// TIA Portal project "Catalyst_syzygy_v2.1" (V17) (continued)
VERSION : 1.0
// stored: InstanceOfName TX-AI
"TX-AI"
BEGIN
   Retain.HMI.Config.ESMXV := 50.0;
   Retain.HMI.Config.SP.Limits.H := 10.0;
   Retain.HMI.Config.SP.Limits.HH := 50.0;
END_DATA_BLOCK

// folder: Analogs inputs/Trasmitters/Level Trasmitters/Datablocks

DATA_BLOCK "LT-1011_DB"   // DB8
{ S7_Optimized_Access := 'TRUE' }
VERSION : 1.0
// stored: InstanceOfName TX-AI
"TX-AI"
BEGIN
   Retain.HMI.Config.SP.Limits.H := 85.0;
   Retain.HMI.Config.SP.Limits.HH := 95.0;
END_DATA_BLOCK

DATA_BLOCK "LT-1061_DB"   // DB9
{ S7_Optimized_Access := 'TRUE' }
VERSION : 1.0
// stored: InstanceOfName TX-AI
"TX-AI"
BEGIN
END_DATA_BLOCK

DATA_BLOCK "LT-1021_DB"   // DB35
{ S7_Optimized_Access := 'TRUE' }
VERSION : 1.0
// stored: InstanceOfName TX-AI
"TX-AI"
BEGIN
END_DATA_BLOCK

DATA_BLOCK "LT-2011_DB"   // DB49
{ S7_Optimized_Access := 'TRUE' }
VERSION : 1.0
// stored: InstanceOfName TX-AI
"TX-AI"
BEGIN
   Retain.HMI.Config.SP.Limits.L := 18.0;
END_DATA_BLOCK

DATA_BLOCK "LT-2021_DB"   // DB56
{ S7_Optimized_Access := 'TRUE' }
VERSION : 1.0
// stored: InstanceOfName TX-AI
"TX-AI"
BEGIN
   Retain.HMI.Config.SP.Limits.L := 18.0;
END_DATA_BLOCK

DATA_BLOCK "LT-1031_DB"   // DB60
{ S7_Optimized_Access := 'TRUE' }
VERSION : 1.0
// stored: InstanceOfName TX-AI
"TX-AI"
BEGIN
END_DATA_BLOCK

DATA_BLOCK "LT-1051_DB"   // DB120
{ S7_Optimized_Access := 'TRUE' }
VERSION : 1.0
// stored: InstanceOfName TX-AI
"TX-AI"
BEGIN
END_DATA_BLOCK

DATA_BLOCK "LT-1011_VOL_DB"   // DB152
{ S7_Optimized_Access := 'TRUE' }
VERSION : 1.0
// stored: InstanceOfName TX-AI
"TX-AI"
BEGIN
   Retain.HMI.Config.ESMXV := 1133.72;
   Retain.HMI.Config.SP.Limits.H := 1000.0;
   Retain.HMI.Config.SP.Limits.HH := 1100.0;
END_DATA_BLOCK

DATA_BLOCK "LT-1061_VOL_DB"   // DB232
{ S7_Optimized_Access := 'TRUE' }
VERSION : 1.0
// stored: InstanceOfName TX-AI
"TX-AI"
BEGIN
END_DATA_BLOCK

DATA_BLOCK "LT-1021_VOL_DB"   // DB243
{ S7_Optimized_Access := 'TRUE' }
VERSION : 1.0
// stored: InstanceOfName TX-AI
"TX-AI"
BEGIN
   Retain.HMI.Config.ESMXV := 2300.0;
   Retain.HMI.Config.SP.Limits.H := 2000.0;
   Retain.HMI.Config.SP.Limits.HH := 2100.0;
END_DATA_BLOCK

DATA_BLOCK "LT-1031_VOL_DB"   // DB245
{ S7_Optimized_Access := 'TRUE' }
VERSION : 1.0
// stored: InstanceOfName TX-AI
"TX-AI"
BEGIN
   Retain.HMI.Config.ESMXV := 500.0;
   Retain.HMI.Config.SP.Limits.H := 450.0;
   Retain.HMI.Config.SP.Limits.HH := 480.0;
END_DATA_BLOCK

DATA_BLOCK "LT-1051_VOL_DB"   // DB246
{ S7_Optimized_Access := 'TRUE' }
VERSION : 1.0
// stored: InstanceOfName TX-AI
"TX-AI"
BEGIN
END_DATA_BLOCK

DATA_BLOCK "LT-2011_VOL_DB"   // DB247
{ S7_Optimized_Access := 'TRUE' }
VERSION : 1.0
// stored: InstanceOfName TX-AI
"TX-AI"
BEGIN
   Retain.HMI.Config.ESMXV := 200.0;
   Retain.HMI.Config.SP.Limits.H := 180.0;
   Retain.HMI.Config.SP.Limits.HH := 190.0;
END_DATA_BLOCK

DATA_BLOCK "LT-2021_VOL_DB"   // DB248
{ S7_Optimized_Access := 'TRUE' }
VERSION : 1.0
// stored: InstanceOfName TX-AI
"TX-AI"
BEGIN
   Retain.HMI.Config.ESMXV := 200.0;
   Retain.HMI.Config.SP.Limits.H := 180.0;
   Retain.HMI.Config.SP.Limits.HH := 190.0;
END_DATA_BLOCK

// folder: Analogs inputs/Trasmitters/Ph Trasmitters/Datablocks

DATA_BLOCK "pH-2011_DB"   // DB46
{ S7_Optimized_Access := 'TRUE' }
VERSION : 1.0
// stored: InstanceOfName TX-AI
"TX-AI"
BEGIN
   Retain.HMI.Config.ESMXV := 14.0;
   Retain.HMI.Config.SP.Limits.HH := 12.0;
   Retain.HMI.Config.SP.Limits.H := 10.0;
END_DATA_BLOCK

DATA_BLOCK "pH-2012_DB"   // DB47
{ S7_Optimized_Access := 'TRUE' }
VERSION : 1.0
// stored: InstanceOfName TX-AI
"TX-AI"
BEGIN
   Retain.HMI.Config.ESMXV := 14.0;
   Retain.HMI.Config.SP.Limits.HH := 12.0;
   Retain.HMI.Config.SP.Limits.H := 10.0;
END_DATA_BLOCK

DATA_BLOCK "pH-2021_DB"   // DB54
{ S7_Optimized_Access := 'TRUE' }
VERSION : 1.0
// stored: InstanceOfName TX-AI
"TX-AI"
BEGIN
   Retain.HMI.Config.ESMXV := 14.0;
   Retain.HMI.Config.SP.Limits.HH := 12.0;
   Retain.HMI.Config.SP.Limits.H := 10.0;
END_DATA_BLOCK

DATA_BLOCK "pH-2022_DB"   // DB55
{ S7_Optimized_Access := 'TRUE' }
VERSION : 1.0
// stored: InstanceOfName TX-AI
"TX-AI"
BEGIN
   Retain.HMI.Config.ESMXV := 14.0;
   Retain.HMI.Config.SP.Limits.HH := 12.0;
   Retain.HMI.Config.SP.Limits.H := 10.0;
END_DATA_BLOCK

// folder: Analogs inputs/Trasmitters/Pressure Trasmitters/Datablocks

DATA_BLOCK "PT-101A_DB"   // DB31
{ S7_Optimized_Access := 'TRUE' }
VERSION : 1.0
// stored: InstanceOfName TX-AI
"TX-AI"
BEGIN
   Retain.HMI.Config.SP.Limits.HH := 124.0;
   Retain.HMI.Config.SP.Limits.H := 120.0;
   Retain.HMI.Config.ESMXV := 125.0;
END_DATA_BLOCK

DATA_BLOCK "PT-101B_DB"   // DB32
{ S7_Optimized_Access := 'TRUE' }
VERSION : 1.0
// stored: InstanceOfName TX-AI
"TX-AI"
BEGIN
   Retain.HMI.Config.SP.Limits.HH := 124.0;
   Retain.HMI.Config.SP.Limits.H := 120.0;
   Retain.HMI.Config.ESMXV := 125.0;
END_DATA_BLOCK

DATA_BLOCK "PT-102A_DB"   // DB36
{ S7_Optimized_Access := 'TRUE' }
VERSION : 1.0
// stored: InstanceOfName TX-AI
"TX-AI"
BEGIN
   Retain.HMI.Config.ESMXV := 125.0;
   Retain.HMI.Config.SP.Limits.HH := 124.0;
   Retain.HMI.Config.SP.Limits.H := 120.0;
END_DATA_BLOCK

DATA_BLOCK "PT-102B_DB"   // DB37
{ S7_Optimized_Access := 'TRUE' }
VERSION : 1.0
// stored: InstanceOfName TX-AI
"TX-AI"
BEGIN
   Retain.HMI.Config.ESMXV := 125.0;
   Retain.HMI.Config.SP.Limits.HH := 124.0;
   Retain.HMI.Config.SP.Limits.H := 120.0;
END_DATA_BLOCK

DATA_BLOCK "PT-201A_DB"   // DB50
{ S7_Optimized_Access := 'TRUE' }
VERSION : 1.0
// stored: InstanceOfName TX-AI
"TX-AI"
BEGIN
   Retain.HMI.Config.ESMXV := 125.0;
   Retain.HMI.Config.SP.Limits.HH := 110.0;
   Retain.HMI.Config.SP.Limits.H := 100.0;
END_DATA_BLOCK

DATA_BLOCK "PT-201B_DB"   // DB51
{ S7_Optimized_Access := 'TRUE' }
VERSION : 1.0
// stored: InstanceOfName TX-AI
"TX-AI"
BEGIN
   Retain.HMI.Config.ESMXV := 125.0;
   Retain.HMI.Config.SP.Limits.HH := 110.0;
   Retain.HMI.Config.SP.Limits.H := 100.0;
END_DATA_BLOCK

DATA_BLOCK "PT-202A_DB"   // DB57
{ S7_Optimized_Access := 'TRUE' }
VERSION : 1.0
// stored: InstanceOfName TX-AI
"TX-AI"
BEGIN
   Retain.HMI.Config.ESMXV := 125.0;
   Retain.HMI.Config.SP.Limits.HH := 110.0;
   Retain.HMI.Config.SP.Limits.H := 100.0;
END_DATA_BLOCK

DATA_BLOCK "PT-202B_DB"   // DB58
{ S7_Optimized_Access := 'TRUE' }
VERSION : 1.0
// stored: InstanceOfName TX-AI
"TX-AI"
BEGIN
   Retain.HMI.Config.ESMXV := 125.0;
   Retain.HMI.Config.SP.Limits.HH := 110.0;
   Retain.HMI.Config.SP.Limits.H := 100.0;
END_DATA_BLOCK

DATA_BLOCK "PT-103A_DB"   // DB61
{ S7_Optimized_Access := 'TRUE' }
VERSION : 1.0
// stored: InstanceOfName TX-AI
"TX-AI"
BEGIN
   Retain.HMI.Config.ESMXV := 125.0;
   Retain.HMI.Config.SP.Limits.H := 124.0;
   Retain.HMI.Config.SP.Limits.L := 120.0;
END_DATA_BLOCK

DATA_BLOCK "PT-103B_DB"   // DB62
{ S7_Optimized_Access := 'TRUE' }
VERSION : 1.0
// stored: InstanceOfName TX-AI
"TX-AI"
BEGIN
   Retain.HMI.Config.ESMXV := 125.0;
   Retain.HMI.Config.SP.Limits.HH := 124.0;
   Retain.HMI.Config.SP.Limits.H := 120.0;
END_DATA_BLOCK

DATA_BLOCK "PT-301A_DB"   // DB64
{ S7_Optimized_Access := 'TRUE' }
VERSION : 1.0
// stored: InstanceOfName TX-AI
"TX-AI"
BEGIN
   Retain.HMI.Config.ESMXV := 125.0;
   Retain.HMI.Config.SP.Limits.HH := 110.0;
   Retain.HMI.Config.SP.Limits.H := 100.0;
END_DATA_BLOCK

DATA_BLOCK "PT-301B_DB"   // DB65
{ S7_Optimized_Access := 'TRUE' }
VERSION : 1.0
// stored: InstanceOfName TX-AI
"TX-AI"
BEGIN
   Retain.HMI.Config.ESMXV := 125.0;
   Retain.HMI.Config.SP.Limits.HH := 110.0;
   Retain.HMI.Config.SP.Limits.H := 100.0;
END_DATA_BLOCK

DATA_BLOCK "PT-104A_DB"   // DB124
{ S7_Optimized_Access := 'TRUE' }
VERSION : 1.0
// stored: InstanceOfName TX-AI
"TX-AI"
BEGIN
   Retain.HMI.Config.ESMXV := 64.0;
END_DATA_BLOCK

DATA_BLOCK "PT-104B_DB"   // DB125
{ S7_Optimized_Access := 'TRUE' }
VERSION : 1.0
// stored: InstanceOfName TX-AI
"TX-AI"
BEGIN
   Retain.HMI.Config.ESMXV := 64.0;
END_DATA_BLOCK

DATA_BLOCK "MFC-4011-P_DB"   // DB162
{ S7_Optimized_Access := 'TRUE' }
VERSION : 1.0
// stored: InstanceOfName TX-AI
"TX-AI"
BEGIN
   Retain.HMI.Config.SP.Limits.HH := 17.3;
   Retain.HMI.Config.SP.Limits.H := 16.3;
   Retain.HMI.Config.SP.Limits.L := 15.0;
   Retain.HMI.Config.SP.Limits.LL := 14.8;
   Retain.HMI.Config.PT.HLD.ALL := t#15s;
   Retain.HMI.Config.PT.HLD.AHH := t#15s;
END_DATA_BLOCK

DATA_BLOCK "PT-M_4024_DB"   // DB165
{ S7_Optimized_Access := 'TRUE' }
VERSION : 1.0
// stored: InstanceOfName TX-AI
"TX-AI"
BEGIN
END_DATA_BLOCK

DATA_BLOCK "PT-M_4025_DB"   // DB166
{ S7_Optimized_Access := 'TRUE' }
VERSION : 1.0
// stored: InstanceOfName TX-AI
"TX-AI"
BEGIN
END_DATA_BLOCK

DATA_BLOCK "MFC-4012-P_DB"   // DB176
{ S7_Optimized_Access := 'TRUE' }
VERSION : 1.0
// stored: InstanceOfName TX-AI
"TX-AI"
BEGIN
END_DATA_BLOCK

DATA_BLOCK "MFC-4024-P_DB"   // DB213
{ S7_Optimized_Access := 'TRUE' }
VERSION : 1.0
// stored: InstanceOfName TX-AI
"TX-AI"
BEGIN
END_DATA_BLOCK

DATA_BLOCK "MFC-4025-P_DB"   // DB216
{ S7_Optimized_Access := 'TRUE' }
VERSION : 1.0
// stored: InstanceOfName TX-AI
"TX-AI"
BEGIN
END_DATA_BLOCK

DATA_BLOCK "MFC-4021-P_DB"   // DB398
{ S7_Optimized_Access := 'TRUE' }
VERSION : 1.0
// stored: InstanceOfName TX-AI
"TX-AI"
BEGIN
END_DATA_BLOCK

// folder: Analogs inputs/Trasmitters/Temperature Trasmitters/DataBlocks

DATA_BLOCK "TT-2011_DB"   // DB44
{ S7_Optimized_Access := 'TRUE' }
VERSION : 1.0
// stored: InstanceOfName TX-AI
"TX-AI"
BEGIN
   Retain.HMI.Config.SP.Limits.L := 75.0;
   Retain.HMI.Config.SP.Limits.LL := 70.0;
   Retain.HMI.Config.ESMXV := 200.0;
END_DATA_BLOCK

DATA_BLOCK "TT-2012_DB"   // DB45
{ S7_Optimized_Access := 'TRUE' }
VERSION : 1.0
// stored: InstanceOfName TX-AI
"TX-AI"
BEGIN
   Retain.HMI.Config.SP.Limits.L := 75.0;
   Retain.HMI.Config.SP.Limits.LL := 70.0;
   Retain.HMI.Config.ESMXV := 200.0;
END_DATA_BLOCK

DATA_BLOCK "TT-2021_DB"   // DB52
{ S7_Optimized_Access := 'TRUE' }
VERSION : 1.0
// stored: InstanceOfName TX-AI
"TX-AI"
BEGIN
   Retain.HMI.Config.ESMXV := 200.0;
   Retain.HMI.Config.SP.Limits.L := 70.0;
   Retain.HMI.Config.SP.Limits.LL := 75.0;
END_DATA_BLOCK

DATA_BLOCK "TT-2022_DB"   // DB53
{ S7_Optimized_Access := 'TRUE' }
VERSION : 1.0
// stored: InstanceOfName TX-AI
"TX-AI"
BEGIN
   Retain.HMI.Config.SP.Limits.L := 75.0;
   Retain.HMI.Config.SP.Limits.LL := 70.0;
   Retain.HMI.Config.ESMXV := 200.0;
END_DATA_BLOCK

DATA_BLOCK "TT-1031_DB"   // DB59
{ S7_Optimized_Access := 'TRUE' }
VERSION : 1.0
// stored: InstanceOfName TX-AI
"TX-AI"
BEGIN
   Retain.HMI.Config.ESMXV := 200.0;
END_DATA_BLOCK

DATA_BLOCK "TT-401A_DB"   // DB69
{ S7_Optimized_Access := 'TRUE' }
VERSION : 1.0
// stored: InstanceOfName TX-AI
"TX-AI"
BEGIN
   Retain.HMI.Config.ESMXV := 1350.0;
   Retain.HMI.Config.RIMXV := 13500.0;
   Retain.HMI.Config.SP.Limits.HH := 800.0;
   Retain.HMI.Config.SP.Limits.H := 750.0;
END_DATA_BLOCK

DATA_BLOCK "TT-401B_DB"   // DB70
{ S7_Optimized_Access := 'TRUE' }
VERSION : 1.0
// stored: InstanceOfName TX-AI
"TX-AI"
BEGIN
   Retain.HMI.Config.ESMXV := 1350.0;
   Retain.HMI.Config.RIMXV := 13500.0;
   Retain.HMI.Config.SP.Limits.HH := 800.0;
   Retain.HMI.Config.SP.Limits.H := 750.0;
END_DATA_BLOCK

DATA_BLOCK "TT-401C_DB"   // DB71
{ S7_Optimized_Access := 'TRUE' }
VERSION : 1.0
// stored: InstanceOfName TX-AI
"TX-AI"
BEGIN
   Retain.HMI.Config.ESMXV := 1350.0;
   Retain.HMI.Config.RIMXV := 13500.0;
   Retain.HMI.Config.SP.Limits.HH := 800.0;
   Retain.HMI.Config.SP.Limits.H := 750.0;
END_DATA_BLOCK

DATA_BLOCK "TT-PT-100_DB"   // DB121
{ S7_Optimized_Access := 'TRUE' }
VERSION : 1.0
// stored: InstanceOfName TX-AI
"TX-AI"
BEGIN
END_DATA_BLOCK

DATA_BLOCK "TE-H201_DB"   // DB128
{ S7_Optimized_Access := 'TRUE' }
VERSION : 1.0
// stored: InstanceOfName TX-AI
"TX-AI"
BEGIN
END_DATA_BLOCK

DATA_BLOCK "TT-4021_DB"   // DB129
{ S7_Optimized_Access := 'TRUE' }
VERSION : 1.0
// stored: InstanceOfName TX-AI
"TX-AI"
BEGIN
END_DATA_BLOCK

DATA_BLOCK "MFC-4011-T_DB"   // DB163
{ S7_Optimized_Access := 'TRUE' }
VERSION : 1.0
// stored: InstanceOfName TX-AI
"TX-AI"
BEGIN
END_DATA_BLOCK

DATA_BLOCK "TE-402A_DB"   // DB209
{ S7_Optimized_Access := 'TRUE' }
VERSION : 1.0
// stored: InstanceOfName TX-AI
"TX-AI"
BEGIN
   Retain.HMI.Config.ESMXV := 1350.0;
   Retain.HMI.Config.RIMXV := 13500.0;
   Retain.HMI.Config.SP.Limits.H := 400.0;
   Retain.HMI.Config.SP.Limits.HH := 480.0;
END_DATA_BLOCK

DATA_BLOCK "TE-402B_DB"   // DB210
{ S7_Optimized_Access := 'TRUE' }
VERSION : 1.0
// stored: InstanceOfName TX-AI
"TX-AI"
BEGIN
   Retain.HMI.Config.ESMXV := 1350.0;
   Retain.HMI.Config.RIMXV := 13500.0;
   Retain.HMI.Config.SP.Limits.HH := 480.0;
   Retain.HMI.Config.SP.Limits.H := 400.0;
END_DATA_BLOCK

DATA_BLOCK "MFC-4024-T_DB"   // DB214
{ S7_Optimized_Access := 'TRUE' }
VERSION : 1.0
// stored: InstanceOfName TX-AI
"TX-AI"
BEGIN
END_DATA_BLOCK

DATA_BLOCK "MFC-4025-T_DB"   // DB217
{ S7_Optimized_Access := 'TRUE' }
VERSION : 1.0
// stored: InstanceOfName TX-AI
"TX-AI"
BEGIN
END_DATA_BLOCK

DATA_BLOCK "PV-HFC-201_DB"   // DB219
{ S7_Optimized_Access := 'TRUE' }
VERSION : 1.0
// stored: InstanceOfName TX-AI
"TX-AI"
BEGIN
END_DATA_BLOCK

DATA_BLOCK "TE-402C_DB"   // DB228
{ S7_Optimized_Access := 'TRUE' }
VERSION : 1.0
// stored: InstanceOfName TX-AI
"TX-AI"
BEGIN
   Retain.HMI.Config.ESMXV := 1350.0;
   Retain.HMI.Config.RIMXV := 13500.0;
   Retain.HMI.Config.SP.Limits.HH := 480.0;
   Retain.HMI.Config.SP.Limits.H := 400.0;
END_DATA_BLOCK

DATA_BLOCK "TE-402D_DB"   // DB229
{ S7_Optimized_Access := 'TRUE' }
VERSION : 1.0
// stored: InstanceOfName TX-AI
"TX-AI"
BEGIN
   Retain.HMI.Config.ESMXV := 1350.0;
   Retain.HMI.Config.RIMXV := 13500.0;
   Retain.HMI.Config.SP.Limits.HH := 480.0;
   Retain.HMI.Config.SP.Limits.H := 400.0;
END_DATA_BLOCK

DATA_BLOCK "TE-402E_DB"   // DB230
{ S7_Optimized_Access := 'TRUE' }
VERSION : 1.0
// stored: InstanceOfName TX-AI
"TX-AI"
BEGIN
   Retain.HMI.Config.ESMXV := 1350.0;
   Retain.HMI.Config.RIMXV := 13500.0;
   Retain.HMI.Config.SP.Limits.HH := 480.0;
   Retain.HMI.Config.SP.Limits.H := 400.0;
END_DATA_BLOCK

DATA_BLOCK "TT-401D_DB"   // DB231
{ S7_Optimized_Access := 'TRUE' }
VERSION : 1.0
// stored: InstanceOfName TX-AI
"TX-AI"
BEGIN
   Retain.HMI.Config.ESMXV := 1350.0;
   Retain.HMI.Config.RIMXV := 13500.0;
   Retain.HMI.Config.SP.Limits.HH := 800.0;
   Retain.HMI.Config.SP.Limits.H := 750.0;
END_DATA_BLOCK

DATA_BLOCK "TT-H201_DB"   // DB249
{ S7_Optimized_Access := 'TRUE' }
VERSION : 1.0
// stored: InstanceOfName TX-AI
"TX-AI"
BEGIN
END_DATA_BLOCK

DATA_BLOCK "MFC-4012-T_DB"   // DB276
{ S7_Optimized_Access := 'TRUE' }
VERSION : 1.0
// stored: InstanceOfName TX-AI
"TX-AI"
BEGIN
END_DATA_BLOCK

DATA_BLOCK "TT-2012B_DB"   // DB372
{ S7_Optimized_Access := 'TRUE' }
VERSION : 1.0
// stored: InstanceOfName TX-AI
"TX-AI"
BEGIN
END_DATA_BLOCK

DATA_BLOCK "TT-2011B_DB"   // DB373
{ S7_Optimized_Access := 'TRUE' }
VERSION : 1.0
// stored: InstanceOfName TX-AI
"TX-AI"
BEGIN
END_DATA_BLOCK

DATA_BLOCK "TT-2021B_DB"   // DB374
{ S7_Optimized_Access := 'TRUE' }
VERSION : 1.0
// stored: InstanceOfName TX-AI
"TX-AI"
BEGIN
END_DATA_BLOCK

DATA_BLOCK "TT-2022B_DB"   // DB375
{ S7_Optimized_Access := 'TRUE' }
VERSION : 1.0
// stored: InstanceOfName TX-AI
"TX-AI"
BEGIN
END_DATA_BLOCK

DATA_BLOCK "TT-104AC_DB"   // DB384
{ S7_Optimized_Access := 'TRUE' }
VERSION : 1.0
// stored: InstanceOfName TX-AI
"TX-AI"
BEGIN
END_DATA_BLOCK

DATA_BLOCK "TT-104BC_DB"   // DB385
{ S7_Optimized_Access := 'TRUE' }
VERSION : 1.0
// stored: InstanceOfName TX-AI
"TX-AI"
BEGIN
END_DATA_BLOCK

DATA_BLOCK "TT-104CC_DB"   // DB386
{ S7_Optimized_Access := 'TRUE' }
VERSION : 1.0
// stored: InstanceOfName TX-AI
"TX-AI"
BEGIN
END_DATA_BLOCK

DATA_BLOCK "MFC-4021-T_DB"   // DB415
{ S7_Optimized_Access := 'TRUE' }
VERSION : 1.0
// stored: InstanceOfName TX-AI
"TX-AI"
BEGIN
END_DATA_BLOCK

// folder: Analogs inputs/Trasmitters/Temperature Trasmitters/Temperature Voting Datablocks

DATA_BLOCK "TT-401 Analog Voting_DB"   // DB146
{ S7_Optimized_Access := 'TRUE' }
VERSION : 0.1
// stored: InstanceOfName 3 Analog Voting
"3 Analog Voting"
BEGIN
END_DATA_BLOCK

DATA_BLOCK "TT-402 Analog Voting_DB"   // DB250
{ S7_Optimized_Access := 'TRUE' }
VERSION : 0.1
// stored: InstanceOfName 3 Analog Voting
"3 Analog Voting"
BEGIN
END_DATA_BLOCK

// folder: Analogs inputs/Trasmitters/VFD_Feedback Trasmitters/Datablocks

DATA_BLOCK "ZT-T101_DB"   // DB72
{ S7_Optimized_Access := 'TRUE' }
VERSION : 1.0
// stored: InstanceOfName TX-AI
"TX-AI"
BEGIN
   Retain.HMI.Config.SP.Limits.H := 90.0;
   Retain.HMI.Config.SP.Limits.HH := 93.0;
END_DATA_BLOCK

DATA_BLOCK "ZT-T102_DB"   // DB73
{ S7_Optimized_Access := 'TRUE' }
VERSION : 1.0
// stored: InstanceOfName TX-AI
"TX-AI"
BEGIN
   Retain.HMI.Config.SP.Limits.H := 90.0;
   Retain.HMI.Config.SP.Limits.HH := 93.0;
END_DATA_BLOCK

DATA_BLOCK "ZT-R201_DB"   // DB74
{ S7_Optimized_Access := 'TRUE' }
VERSION : 1.0
// stored: InstanceOfName TX-AI
"TX-AI"
BEGIN
END_DATA_BLOCK

DATA_BLOCK "ZT-R202_DB"   // DB75
{ S7_Optimized_Access := 'TRUE' }
VERSION : 1.0
// stored: InstanceOfName TX-AI
"TX-AI"
BEGIN
END_DATA_BLOCK

DATA_BLOCK "ZT-C301_DB"   // DB402
{ S7_Optimized_Access := 'TRUE' }
VERSION : 1.0
// stored: InstanceOfName TX-AI
"TX-AI"
BEGIN
   Retain.HMI.Config.ESMXV := 1750.0;
END_DATA_BLOCK

// folder: Analogs inputs/Trasmitters/Vibration Transmitter

DATA_BLOCK "VT-C301_DB"   // DB168
{ S7_Optimized_Access := 'TRUE' }
VERSION : 1.0
// stored: InstanceOfName TX-AI
"TX-AI"
BEGIN
   Retain.HMI.Config.ESMXV := 50.0;
   Retain.HMI.Config.SP.Limits.H := 30.0;
   Retain.HMI.Config.SP.Limits.HH := 37.5;
END_DATA_BLOCK

// folder: Analogs inputs/Trasmitters/average

DATA_BLOCK "TT-R-201_Average_DB"   // DB170
{ S7_Optimized_Access := 'TRUE' }
VERSION : 0.1
// stored: InstanceOfName Average
"Average"
BEGIN
END_DATA_BLOCK

DATA_BLOCK "TT-R-202_Average_DB"   // DB171
{ S7_Optimized_Access := 'TRUE' }
VERSION : 0.1
// stored: InstanceOfName Average
"Average"
BEGIN
END_DATA_BLOCK

DATA_BLOCK "TT-R-201/R-202_Average_DB"   // DB172
{ S7_Optimized_Access := 'TRUE' }
VERSION : 0.1
// stored: InstanceOfName Average
"Average"
BEGIN
END_DATA_BLOCK

DATA_BLOCK "PH-R-201_Average_DB"   // DB220
{ S7_Optimized_Access := 'TRUE' }
VERSION : 0.1
// stored: InstanceOfName Average
"Average"
BEGIN
END_DATA_BLOCK

DATA_BLOCK "PH-R-202_Average_DB"   // DB221
{ S7_Optimized_Access := 'TRUE' }
VERSION : 0.1
// stored: InstanceOfName Average
"Average"
BEGIN
END_DATA_BLOCK

DATA_BLOCK "PH-R-201/R-202_Average_DB"   // DB222
{ S7_Optimized_Access := 'TRUE' }
VERSION : 0.1
// stored: InstanceOfName Average
"Average"
BEGIN
END_DATA_BLOCK

// folder: Calculations

DATA_BLOCK "TC-R402A_Ramp_DB"   // DB157
{ S7_Optimized_Access := 'TRUE' }
VERSION : 0.1
// stored: InstanceOfName Ramp_v2
"Ramp_v2"
BEGIN
END_DATA_BLOCK

DATA_BLOCK "TC-R402B_Ramp_DB"   // DB158
{ S7_Optimized_Access := 'TRUE' }
VERSION : 0.1
// stored: InstanceOfName Ramp_v2
"Ramp_v2"
BEGIN
END_DATA_BLOCK

// folder: Cause&EffectMatrix

DATA_BLOCK "CEM1_DB"   // DB90
{ S7_Optimized_Access := 'TRUE' }
VERSION : 0.1
// stored: InstanceOfName CauseAndEffect
"CauseAndEffect"
BEGIN
END_DATA_BLOCK

// folder: Diagnostic

DATA_BLOCK "Diag_DB"   // DB89
{ S7_Optimized_Access := 'TRUE' }
VERSION : 0.1
// stored: InstanceOfName diag
"diag"
BEGIN
END_DATA_BLOCK

// folder: ESD

DATA_BLOCK "R-201_Interlocks_DB"   // DB267
{ S7_Optimized_Access := 'TRUE' }
VERSION : 0.1
// stored: InstanceOfName Interlocks
"Interlocks"
BEGIN
END_DATA_BLOCK

DATA_BLOCK "T-104_Interlocks_DB"   // DB346
{ S7_Optimized_Access := 'TRUE' }
VERSION : 0.1
// stored: InstanceOfName Interlocks
"Interlocks"
BEGIN
END_DATA_BLOCK

DATA_BLOCK "R-202_Interlocks_DB"   // DB347
{ S7_Optimized_Access := 'TRUE' }
VERSION : 0.1
// stored: InstanceOfName Interlocks
"Interlocks"
BEGIN
END_DATA_BLOCK

DATA_BLOCK "T-101_Interlocks_DB"   // DB348
{ S7_Optimized_Access := 'TRUE' }
VERSION : 0.1
// stored: InstanceOfName Interlocks
"Interlocks"
BEGIN
END_DATA_BLOCK

DATA_BLOCK "T-102_Interlocks_DB"   // DB349
{ S7_Optimized_Access := 'TRUE' }
VERSION : 0.1
// stored: InstanceOfName Interlocks
"Interlocks"
BEGIN
END_DATA_BLOCK

DATA_BLOCK "T-103_Interlocks_DB"   // DB350
{ S7_Optimized_Access := 'TRUE' }
VERSION : 0.1
// stored: InstanceOfName Interlocks
"Interlocks"
BEGIN
END_DATA_BLOCK

DATA_BLOCK "Centrifuge_Interlocks_DB"   // DB351
{ S7_Optimized_Access := 'TRUE' }
VERSION : 0.1
// stored: InstanceOfName Interlocks
"Interlocks"
BEGIN
END_DATA_BLOCK

// folder: ESD/Datablocks/C-301

DATA_BLOCK "C-301 Centrifuge_INTERLOCKS"   // DB193
{ S7_Optimized_Access := 'TRUE' }
VERSION : 0.1
// stored: InstanceOfName Interlocks
"Interlocks"
BEGIN
END_DATA_BLOCK

// folder: ESD/Datablocks/H-401

DATA_BLOCK "I401_Calcination_Interlocks"   // DB211
{ S7_Optimized_Access := 'TRUE' }
VERSION : 0.1
// stored: InstanceOfName Interlocks
"Interlocks"
BEGIN
END_DATA_BLOCK

// folder: ESD/Datablocks/H-402

DATA_BLOCK "I402_Passivate_Interlocks"   // DB192
{ S7_Optimized_Access := 'TRUE' }
VERSION : 0.1
// stored: InstanceOfName Interlocks
"Interlocks"
BEGIN
END_DATA_BLOCK

// folder: ESD/Datablocks/R-201

DATA_BLOCK "I201A_Reactor_Interlocks"   // DB195
{ S7_Optimized_Access := 'TRUE' }
VERSION : 0.1
// stored: InstanceOfName Interlocks
"Interlocks"
BEGIN
END_DATA_BLOCK

DATA_BLOCK "I201B_Reactor_Interlocks"   // DB197
{ S7_Optimized_Access := 'TRUE' }
VERSION : 0.1
// stored: InstanceOfName Interlocks
"Interlocks"
BEGIN
END_DATA_BLOCK

// folder: ESD/Datablocks/R-202

DATA_BLOCK "I202A_Reactors_Interlocks"   // DB196
{ S7_Optimized_Access := 'TRUE' }
VERSION : 0.1
// stored: InstanceOfName Interlocks
"Interlocks"
BEGIN
END_DATA_BLOCK

DATA_BLOCK "I202B_Reactors_Interlocks"   // DB198
{ S7_Optimized_Access := 'TRUE' }
VERSION : 0.1
// stored: InstanceOfName Interlocks
"Interlocks"
BEGIN
END_DATA_BLOCK

// folder: ESD/Datablocks/T-101

DATA_BLOCK "T-101 Mix & Wash X material INTERLOCKS"   // DB233
{ S7_Optimized_Access := 'TRUE' }
VERSION : 0.1
// stored: InstanceOfName Interlocks
"Interlocks"
BEGIN
END_DATA_BLOCK

// folder: ESD/Datablocks/T-102

DATA_BLOCK "T-102 Mix & Wash Y Material  INTERLOCKS"   // DB194
{ S7_Optimized_Access := 'TRUE' }
VERSION : 0.1
// stored: InstanceOfName Interlocks
"Interlocks"
BEGIN
   HMI.Bypass_1 := true;
   HMI.Bypass_2 := true;
   HMI.Bypass_3 := true;
   HMI.Bypass_4 := true;
   HMI.Bypass_5 := true;
   HMI.Bypass_7 := true;
   HMI.Bypass_6 := true;
   HMI.Bypass_8 := true;
   HMI.Bypass_9 := true;
   HMI.Bypass_10 := true;
   HMI.Bypass_11 := true;
   HMI.Bypass_12 := true;
   HMI.Bypass_13 := true;
   HMI.Bypass_14 := true;
   HMI.Bypass_15 := true;
   HMI.Bypass_16 := true;
   HMI.Bypass_17 := true;
   HMI.Bypass_18 := true;
   HMI.Bypass_19 := true;
   HMI.Bypass_20 := true;
   HMI.Bypass_21 := true;
   HMI.Bypass_22 := true;
   HMI.Bypass_23 := true;
   HMI.Bypass_24 := true;
   HMI.Bypass_25 := true;
   HMI.Bypass_26 := true;
   HMI.Bypass_27 := true;
   HMI.Bypass_28 := true;
   HMI.Bypass_29 := true;
   HMI.Bypass_30 := true;
   HMI.Bypass_31 := true;
   HMI.Bypass_32 := true;
END_DATA_BLOCK

// folder: ESD/Datablocks/T-103

DATA_BLOCK "I103A_Reactor_Interlocks"   // DB205
{ S7_Optimized_Access := 'TRUE' }
VERSION : 0.1
// stored: InstanceOfName Interlocks
"Interlocks"
BEGIN
END_DATA_BLOCK

DATA_BLOCK "I103B_Reactor_Interlocks"   // DB206
{ S7_Optimized_Access := 'TRUE' }
VERSION : 0.1
// stored: InstanceOfName Interlocks
"Interlocks"
BEGIN
END_DATA_BLOCK

DATA_BLOCK "I103C_Reactor_Interlocks"   // DB207
{ S7_Optimized_Access := 'TRUE' }
VERSION : 0.1
// stored: InstanceOfName Interlocks
"Interlocks"
BEGIN
END_DATA_BLOCK

DATA_BLOCK "I103D_Reactor_Interlocks"   // DB208
{ S7_Optimized_Access := 'TRUE' }
VERSION : 0.1
// stored: InstanceOfName Interlocks
"Interlocks"
BEGIN
END_DATA_BLOCK

// folder: Outside Comms/Centrifuge

DATA_BLOCK "ExchangeCentrifuge_DB"   // DB265
{ S7_Optimized_Access := 'TRUE' }
VERSION : 0.1
   VAR
      ToCentrifuge : Struct
         SS : Bool;   // Start/Stop Command
         "E-Stop" : Bool;   // Emergency Stop to Centrifuge from DCS
         Reset : Bool;   // Ret. Feeler and Fault Reset
         FeelerEngage : Bool;   // Feeler Engage
         SP : Int;   // Centrifuge Speed Setpoint
      END_STRUCT;
      FromCentrifuge : Struct
         VibFault : Bool;   // Vibration Fault
         "E-Stop" : Bool;   // Emergency Stop to DCS from Centrifuge
         S_Fault : Bool;   // System Fault
         BsktFull : Bool;   // Centrifuge Basket Full
         CoverNLock : Bool;   // Centrifuge Cover Not Locked
         FeelerRetracted : Bool;   // Centrifuge Feeler Retracted
         "VT-8" : Int;   // Vibration Transmitter
         PV : Int;   // Centrifuge Speed Feedback
      END_STRUCT;
   END_VAR
BEGIN
END_DATA_BLOCK

// folder: Outside Comms/ModBus Comms/CO/CO2/O2 R-401 Analizer

DATA_BLOCK "COCO2O_R-401_MB_rDT_DB"   // DB159
{ S7_Optimized_Access := 'TRUE' }
AUTHOR : JL
VERSION : 0.1
// stored: InstanceOfName MFC_MB_rDT
"MFC_MB_rDT"
BEGIN
END_DATA_BLOCK

DATA_BLOCK "COCO2O_R401_MB_iDT_DB"   // DB242
{ S7_Optimized_Access := 'TRUE' }
AUTHOR : JL
VERSION : 0.1
// stored: InstanceOfName MFC_MB_iDT
"MFC_MB_iDT"
BEGIN
END_DATA_BLOCK

DATA_BLOCK "COCO2O_MB_ByteDT_DB"   // DB275
{ S7_Optimized_Access := 'TRUE' }
AUTHOR : JL
VERSION : 0.1
// stored: InstanceOfName MFC_MB_ByteDT
"MFC_MB_ByteDT"
BEGIN
END_DATA_BLOCK

DATA_BLOCK "test_Tcon"   // DB278
{ S7_Optimized_Access := 'TRUE' }
VERSION : 0.1
   VAR
      connects : TCON_IP_v4;
   END_VAR
BEGIN
   connects.InterfaceId := 258;
   connects.ID := 39;
   connects.RemotePort := 502;
   connects.RemoteAddress.ADDR[1] := 192;
   connects.RemoteAddress.ADDR[2] := 168;
   connects.RemoteAddress.ADDR[3] := 2;
   connects.RemoteAddress.ADDR[4] := 32;
END_DATA_BLOCK

// folder: Outside Comms/ModBus Comms/EurothermControllers

DATA_BLOCK "Eurothem_Data"   // DB251
{ S7_Optimized_Access := 'TRUE' }
VERSION : 0.1
   VAR
      Read : Struct
         Read1 : "ModBus_Data";
         Read2 : "ModBus_Data";
         Read3 : "ModBus_Data";
      END_STRUCT;
      Write : Struct
         Write1 : "ModBus_Data";   // Write from address 40023
         Write2 : "ModBus_Data";   // Write from address 41280
      END_STRUCT;
   END_VAR
BEGIN
END_DATA_BLOCK

// folder: Outside Comms/ModBus Comms/EurothermControllers/TC-4011A

DATA_BLOCK "TC-4011A_DB"   // DB134
{ S7_Optimized_Access := 'TRUE' }
VERSION : 0.1
   VAR
      Data : "EurothermCtls_UDT";
      AddrCtrl : Struct
         CurrentAddr : UDInt;
         Down : Bool;
         Up : Bool;
         RisingUp : Bool;
      END_STRUCT;
   END_VAR
BEGIN
END_DATA_BLOCK

DATA_BLOCK "TC-4011A_R1"   // DB252
{ S7_Optimized_Access := 'TRUE' }
AUTHOR : JL
VERSION : 0.1
// stored: InstanceOfName Eurotherm_MB_FB
"Eurotherm_MB_FB"
BEGIN
END_DATA_BLOCK

DATA_BLOCK "TC-4011A_R2"   // DB255
{ S7_Optimized_Access := 'TRUE' }
AUTHOR : JL
VERSION : 0.1
// stored: InstanceOfName Eurotherm_MB_FB
"Eurotherm_MB_FB"
BEGIN
END_DATA_BLOCK

DATA_BLOCK "TC-4011A_R3"   // DB256
{ S7_Optimized_Access := 'TRUE' }
AUTHOR : JL
VERSION : 0.1
// stored: InstanceOfName Eurotherm_MB_FB
"Eurotherm_MB_FB"
BEGIN
END_DATA_BLOCK

DATA_BLOCK "TC-4011A_W1"   // DB257
{ S7_Optimized_Access := 'TRUE' }
AUTHOR : JL
VERSION : 0.1
// stored: InstanceOfName Eurotherm_MB_FB
"Eurotherm_MB_FB"
BEGIN
END_DATA_BLOCK

DATA_BLOCK "TC-4011A_W2"   // DB258
{ S7_Optimized_Access := 'TRUE' }
AUTHOR : JL
VERSION : 0.1
// stored: InstanceOfName Eurotherm_MB_FB
"Eurotherm_MB_FB"
BEGIN
END_DATA_BLOCK

DATA_BLOCK "TC-4011A_W3"   // DB259
{ S7_Optimized_Access := 'TRUE' }
AUTHOR : JL
VERSION : 0.1
// stored: InstanceOfName Eurotherm_MB_FB
"Eurotherm_MB_FB"
BEGIN
END_DATA_BLOCK

DATA_BLOCK "TC-4011A_W4"   // DB260
{ S7_Optimized_Access := 'TRUE' }
AUTHOR : JL
VERSION : 0.1
// stored: InstanceOfName Eurotherm_MB_FB
"Eurotherm_MB_FB"
BEGIN
END_DATA_BLOCK

// folder: Outside Comms/ModBus Comms/EurothermControllers/TC-4011B

DATA_BLOCK "TC-4011B_DB"   // DB189
{ S7_Optimized_Access := 'TRUE' }
VERSION : 0.1
   VAR
      Data : "EurothermCtls_UDT";
      MBLogic : Struct
         OS : Array[0..31] of Bool;
      END_STRUCT;
   END_VAR
BEGIN
END_DATA_BLOCK

DATA_BLOCK "TC-4011B_R1"   // DB261
{ S7_Optimized_Access := 'TRUE' }
AUTHOR : JL
VERSION : 0.1
// stored: InstanceOfName Eurotherm_MB_FB
"Eurotherm_MB_FB"
BEGIN
END_DATA_BLOCK

DATA_BLOCK "TC-4011B_R2"   // DB382
{ S7_Optimized_Access := 'TRUE' }
AUTHOR : JL
VERSION : 0.1
// stored: InstanceOfName Eurotherm_MB_FB
"Eurotherm_MB_FB"
BEGIN
END_DATA_BLOCK

DATA_BLOCK "TC-4011B_R3"   // DB403
{ S7_Optimized_Access := 'TRUE' }
AUTHOR : JL
VERSION : 0.1
// stored: InstanceOfName Eurotherm_MB_FB
"Eurotherm_MB_FB"
BEGIN
END_DATA_BLOCK

DATA_BLOCK "TC-4011B_W1"   // DB406
{ S7_Optimized_Access := 'TRUE' }
AUTHOR : JL
VERSION : 0.1
// stored: InstanceOfName Eurotherm_MB_FB
"Eurotherm_MB_FB"
BEGIN
END_DATA_BLOCK

DATA_BLOCK "TC-4011B_W2"   // DB408
{ S7_Optimized_Access := 'TRUE' }
AUTHOR : JL
VERSION : 0.1
// stored: InstanceOfName Eurotherm_MB_FB
"Eurotherm_MB_FB"
BEGIN
END_DATA_BLOCK

DATA_BLOCK "TC-4011B_W3"   // DB409
{ S7_Optimized_Access := 'TRUE' }
AUTHOR : JL
VERSION : 0.1
// stored: InstanceOfName Eurotherm_MB_FB
"Eurotherm_MB_FB"
BEGIN
END_DATA_BLOCK

DATA_BLOCK "TC-4011B_W4"   // DB412
{ S7_Optimized_Access := 'TRUE' }
AUTHOR : JL
VERSION : 0.1
// stored: InstanceOfName Eurotherm_MB_FB
"Eurotherm_MB_FB"
BEGIN
END_DATA_BLOCK

// folder: Outside Comms/ModBus Comms/EurothermControllers/TC-4011C

DATA_BLOCK "TC-4011C_DB"   // DB179
{ S7_Optimized_Access := 'TRUE' }
VERSION : 0.1
   VAR
      Data : "EurothermCtls_UDT";
      MBLogic : Struct
         ResetErrors : Bool;
         Start : Bool;
         ReStart : Bool;
         R1_Ready : Bool;
         R1_Processing : Bool;
         R1_Done : Bool;
         R2_Ready : Bool;
         R2_Processing : Bool;
         R2_Done : Bool;
         R3_Ready : Bool;
         R3_Processing : Bool;
         R3_Done : Bool;
         W1_Ready : Bool;
         W1_Processing : Bool;
         W1_Done : Bool;
         W2_Ready : Bool;
         W2_Processing : Bool;
         W2_Done : Bool;
         DoneCtrl : Struct
            R1_Dn : Bool;
            R2_Dn : Bool;
            R3_Dn : Bool;
            W1_Dn : Bool;
            W2_Dn : Bool;
         END_STRUCT;
         SelectorToRead : Array[0..31] of Bool;
      END_STRUCT;
   END_VAR
BEGIN
END_DATA_BLOCK

DATA_BLOCK "TC-4011C_R1"   // DB262
{ S7_Optimized_Access := 'TRUE' }
AUTHOR : JL
VERSION : 0.1
// stored: InstanceOfName Eurotherm_MB_FB
"Eurotherm_MB_FB"
BEGIN
END_DATA_BLOCK

DATA_BLOCK "TC-4011C_R2"   // DB383
{ S7_Optimized_Access := 'TRUE' }
AUTHOR : JL
VERSION : 0.1
// stored: InstanceOfName Eurotherm_MB_FB
"Eurotherm_MB_FB"
BEGIN
END_DATA_BLOCK

DATA_BLOCK "TC-4011C_R3"   // DB404
{ S7_Optimized_Access := 'TRUE' }
AUTHOR : JL
VERSION : 0.1
// stored: InstanceOfName Eurotherm_MB_FB
"Eurotherm_MB_FB"
BEGIN
END_DATA_BLOCK

DATA_BLOCK "TC-4011C_W1"   // DB405
{ S7_Optimized_Access := 'TRUE' }
AUTHOR : JL
VERSION : 0.1
// stored: InstanceOfName Eurotherm_MB_FB
"Eurotherm_MB_FB"
BEGIN
END_DATA_BLOCK

DATA_BLOCK "TC-4011C_W2"   // DB407
{ S7_Optimized_Access := 'TRUE' }
AUTHOR : JL
VERSION : 0.1
// stored: InstanceOfName Eurotherm_MB_FB
"Eurotherm_MB_FB"
BEGIN
END_DATA_BLOCK

DATA_BLOCK "TC-4011C_W3"   // DB410
{ S7_Optimized_Access := 'TRUE' }
AUTHOR : JL
VERSION : 0.1
// stored: InstanceOfName Eurotherm_MB_FB
"Eurotherm_MB_FB"
BEGIN
END_DATA_BLOCK

DATA_BLOCK "TC-4011C_W4"   // DB411
{ S7_Optimized_Access := 'TRUE' }
AUTHOR : JL
VERSION : 0.1
// stored: InstanceOfName Eurotherm_MB_FB
"Eurotherm_MB_FB"
BEGIN
END_DATA_BLOCK

// folder: Outside Comms/ModBus Comms/Funace_R-402/TC-402A

DATA_BLOCK "TC-402A_MB_DB"   // DB119
{ S7_Optimized_Access := 'TRUE' }
AUTHOR : JL
VERSION : 0.1
// stored: InstanceOfName YUDIAN_MB_FB
"YUDIAN_MB_FB"
BEGIN
END_DATA_BLOCK

DATA_BLOCK "TC-402A_DB"   // DB424
{ S7_Optimized_Access := 'TRUE' }
VERSION : 0.1
   VAR
      Data : "EurothermCtls_UDT";
      AddrCtrl : Struct
         CurrentAddr : UDInt;
         Down : Bool;
         Up : Bool;
         RisingUp : Bool;
      END_STRUCT;
   END_VAR
BEGIN
END_DATA_BLOCK

DATA_BLOCK "TC-402A_R1"   // DB428
{ S7_Optimized_Access := 'TRUE' }
AUTHOR : JL
VERSION : 0.1
// stored: InstanceOfName Eurotherm_MB_FB
"Eurotherm_MB_FB"
BEGIN
END_DATA_BLOCK

DATA_BLOCK "TC-402A_R2"   // DB430
{ S7_Optimized_Access := 'TRUE' }
AUTHOR : JL
VERSION : 0.1
// stored: InstanceOfName Eurotherm_MB_FB
"Eurotherm_MB_FB"
BEGIN
END_DATA_BLOCK

DATA_BLOCK "TC-402A_R3"   // DB433
{ S7_Optimized_Access := 'TRUE' }
AUTHOR : JL
VERSION : 0.1
// stored: InstanceOfName Eurotherm_MB_FB
"Eurotherm_MB_FB"
BEGIN
END_DATA_BLOCK

DATA_BLOCK "TC-402A_W1"   // DB434
{ S7_Optimized_Access := 'TRUE' }
AUTHOR : JL
VERSION : 0.1
// stored: InstanceOfName Eurotherm_MB_FB
"Eurotherm_MB_FB"
BEGIN
END_DATA_BLOCK

// folder: Outside Comms/ModBus Comms/Funace_R-402/TC-402A/MB_Server

DATA_BLOCK "Data_MB_Server"   // DB148
{ S7_Optimized_Access := 'FALSE' }
VERSION : 0.1
   VAR
      Data : Struct
         fromCtrl : Array[0..124] of Int;
      END_STRUCT;
   END_VAR
BEGIN
END_DATA_BLOCK

// folder: Outside Comms/ModBus Comms/Funace_R-402/TC-402B

DATA_BLOCK "MB_Server_Config"   // DB147
{ S7_Optimized_Access := 'TRUE' }